   "Carrier_63_G120DControlWord.2" AT %I3510.2 : Bool;   // Bit_02_AUS3_STOP
   "Carrier_63_G120DControlWord.3" AT %I3510.3 : Bool;   // Bit_03_EN
   "Carrier_63_G120DControlWord.4" AT %I3510.4 : Bool;   // Bit_04_EN_RAMP
   "Carrier_63_G120DControlWord.5" AT %I3510.5 : Bool;   // Bit_05_START_RAMP
   "Carrier_63_G120DControlWord.6" AT %I3510.6 : Bool;   // Bit_06_SETPOINT
   "Carrier_63_G120DControlWord.7" AT %I3510.7 : Bool;   // Bit_07_RESET
   "Carrier_63_G120DControlWord.8" AT %I3511.0 : Bool;   // Bit_08_JOG_R
   "Carrier_63_G120DControlWord.9" AT %I3511.1 : Bool;   // Bit_09_JOG_L
   "Carrier_63_G120DControlWord.10" AT %I3511.2 : Bool;   // Bit_10_CONTR_PLC
   "Carrier_63_G120DControlWord.11" AT %I3511.3 : Bool;   // Bit_11_REVERSE
   "Carrier_63_G120DControlWord.12" AT %I3511.4 : Bool;   // Bit_12_BRAKE_RELEASE
   "Carrier_63_G120DControlWord.13" AT %I3511.5 : Bool;   // Bit_13_DDS
   "Carrier_63_G120DControlWord.14" AT %I3511.6 : Bool;   // Bit_14_DO0
   "Carrier_63_G120DControlWord.15" AT %I3511.7 : Bool;   // Bit_15_DO1
   "Carrier_63_G120DStatusWord" AT %IW3512 : Word;   // G120D_ZSW1_STATUS
   "Carrier_63_G120DStatusWord.0" AT %I3512.0 : Bool;   // Bit_00_READY_RUN
   "Carrier_63_G120DStatusWord.1" AT %I3512.1 : Bool;   // Bit_01_READY_ON
   "Carrier_63_G120DStatusWord.2" AT %I3512.2 : Bool;   // Bit_02_ENABLE
   "Carrier_63_G120DStatusWord.3" AT %I3512.3 : Bool;   // Bit_03_FAULT
   "Carrier_63_G120DStatusWord.4" AT %I3512.4 : Bool;   // Bit_04_OFF2
   "Carrier_63_G120DStatusWord.5" AT %I3512.5 : Bool;   // Bit_05_OFF3
   "Carrier_63_G120DStatusWord.6" AT %I3512.6 : Bool;   // Bit_06_LOCK_OUT
   "Carrier_63_G120DStatusWord.7" AT %I3512.7 : Bool;   // Bit_07_WARN
   "Carrier_63_G120DStatusWord.8" AT %I3513.0 : Bool;   // Bit_08_NO_DEVIATION
   "Carrier_63_G120DStatusWord.9" AT %I3513.1 : Bool;   // Bit_09_CONTR_PLC
   "Carrier_63_G120DStatusWord.10" AT %I3513.2 : Bool;   // Bit_10_F_MAX
   "Carrier_63_G120DStatusWord.11" AT %I3513.3 : Bool;   // Bit_11_LIMIT_REACHED
   "Carrier_63_G120DStatusWord.12" AT %I3513.4 : Bool;   // Bit_12_BRAKE_OPEN
   "Carrier_63_G120DStatusWord.13" AT %I3513.5 : Bool;   // Bit_13_NO_OVERTEMP
   "Carrier_63_G120DStatusWord.14" AT %I3513.6 : Bool;   // Bit_14_CW_CCW
   "Carrier_63_G120DStatusWord.15" AT %I3513.7 : Bool;   // Bit_15_OVERL
   "Carrier_63_Slot2_Input" AT %IW3514 : Word;   // SLOT 2 INPUT WORD
   "Carrier_63_CrashDetectSW" AT %I3514.0 : Bool;   // CRASH DETECT SW
   "Carrier_63_SpareSafetyInput(2_1)" AT %I3514.1 : Bool;   // SPARE SAFETY INPUT
   "Carrier_63_SpareSafetyInput(2_2)" AT %I3514.2 : Bool;   // SPARE SAFETY INPUT
   "Carrier_63_SpareSafetyInput(2_3)" AT %I3514.3 : Bool;   // SPARE SAFETY INPUT
   "Carrier_63_SpareSafetyInput(2_4)" AT %I3514.4 : Bool;   // SPARE SAFETY INPUT
   "Carrier_63_SpareSafetyInput(2_5)" AT %I3514.5 : Bool;   // SPARE SAFETY INPUT
   "Carrier_63_SpareSafetyInput(2_6)" AT %I3514.6 : Bool;   // SPARE SAFETY INPUT
   "Carrier_63_SpareSafetyInput(2_7)" AT %I3514.7 : Bool;   // SPARE SAFETY INPUT
   "Carrier_63_Slot3_SafetyOutput" AT %IW3515 : Word;   // SLOT 3 SAFETY OUTPUT WORD
   "Carrier_63_Crash_Detect_OK" AT %I3515.0 : Bool;   // CARRIER CRASH DETECT
   "Carrier_63_SpareSafetyOutput(3_1)" AT %I3515.1 : Bool;   // SPARE SAFETY OUTPUT
   "Carrier_63_SpareSafetyOutput(3_2)" AT %I3515.2 : Bool;   // SPARE SAFETY OUTPUT
   "Carrier_63_SpareSafetyOutput(3_3)" AT %I3515.3 : Bool;   // SPARE SAFETY OUTPUT
   "Carrier_63_SpareSafetyOutput(3_4)" AT %I3515.4 : Bool;   // SPARE SAFETY OUTPUT
   "Carrier_63_SpareSafetyOutput(3_5)" AT %I3515.5 : Bool;   // SPARE SAFETY OUTPUT
   "Carrier_63_SpareSafetyOutput(3_6)" AT %I3515.6 : Bool;   // SPARE SAFETY OUTPUT
   "Carrier_63_SpareSafetyOutput(3_7)" AT %I3515.7 : Bool;   // SPARE SAFETY OUTPUT
   "Carrier_63_Slot4_Input" AT %IW3516 : Word;   // SLOT 4 INPUT WORD
   "Carrier_63_480VPowerOn_MDCB1" AT %I3516.0 : Bool;   // 480 VAC POWER ON MDCB 1
   "Carrier_63_SpareInput(4_1)" AT %I3516.1 : Bool;   // SPARE INPUT
   "Carrier_63_SpareInput(4_2)" AT %I3516.2 : Bool;   // SPARE INPUT
   "Carrier_63_SitopSelectStatus" AT %I3516.3 : Bool;   // SITOP SELECT STATUS
   "Carrier_63_DCsupplyOnPSCB2" AT %I3516.4 : Bool;   // DC SUPPLY ON PSCB 2
   "Carrier_63_SpareInput(4_5)" AT %I3516.5 : Bool;   // SPARE INPUT
   "Carrier_63_SpareInput(4_6)" AT %I3516.6 : Bool;   // SPARE INPUT
   "Carrier_63_SpareInput(4_7)" AT %I3516.7 : Bool;   // SPARE INPUT
   "Carrier_63_PB1_ProdHoldLH" AT %I3517.0 : Bool;   // PB 1 PRODUCTION HOLD LH
   "Carrier_63_PB2_ResetLH" AT %I3517.1 : Bool;   // PB 2 RESET LH
   "Carrier_63_PB3_ProdHoldRH" AT %I3517.2 : Bool;   // PB 3 PRODUCTION HOLD RH
   "Carrier_63_PB4_ResetRH" AT %I3517.3 : Bool;   // PB 4 RESET RH
   "Carrier_63_SpareInput(4_14)" AT %I3517.4 : Bool;   // SPARE INPUT
   "Carrier_63_SpareInput(4_15)" AT %I3517.5 : Bool;   // SPARE INPUT
   "Carrier_63_SpareInput(4_16)" AT %I3517.6 : Bool;   // SPARE INPUT
   "Carrier_63_SpareInput(4_17)" AT %I3517.7 : Bool;   // SPARE INPUT
   "Carrier_63_Slot5_Output" AT %IW3518 : Word;   // SLOT 5 OUTPUT WORD
   "Carrier_63_IRD400_HMI_24VDC_ENABLE" AT %I3518.0 : Bool;   // IRD 400 PANEL HMI 24V DC POWER
   "Carrier_63_FaultLight_LH" AT %I3518.1 : Bool;   // FAULT LIGHT LH
   "Carrier_63_RunLight_LH" AT %I3518.2 : Bool;   // RUN LIGHT LH
   "Carrier_63_FaultLight_RH" AT %I3518.3 : Bool;   // FAULT LIGHT RH
   "Carrier_63_RunLight_RH" AT %I3518.4 : Bool;   // RUN LIGHT RH
   "Carrier_63_SpareOutput(5_5)" AT %I3518.5 : Bool;   // SPARE OUTPUT
   "Carrier_63_SpareOutput(5_6)" AT %I3518.6 : Bool;   // SPARE OUTPUT
   "Carrier_63_SpareOutput(5_7)" AT %I3518.7 : Bool;   // SPARE OUTPUT
   "Carrier_63_ActualSpeed" AT %IW3520 : Word;   // ACTUAL SPEED
   "Carrier_63_CarrierDriveAlarm" AT %IW3522 : Word;   // CARRIER DRIVE ALARM
   "Carrier_63_CarrierDriveWarning" AT %IW3524 : Word;   // CARRIER DRIVE WARNING
   "Carrier_64_Status" AT %IW3550 : Word;   // CARRIER STATUS WORD
   "Carrier_64_Status.0" AT %I3550.0 : Bool;   // HEARTBEAT
   "Carrier_64_Status.1" AT %I3550.1 : Bool;   // MANUAL
   "Carrier_64_Status.2" AT %I3550.2 : Bool;   // IN_AUTO
   "Carrier_64_Status.3" AT %I3550.3 : Bool;   // POSITIONING_COMPLETE
   "Carrier_64_Status.4" AT %I3550.4 : Bool;   // PRODUCTION HOLD
   "Carrier_64_Status.5" AT %I3550.5 : Bool;   // CARRIER MOVING FORWARD
   "Carrier_64_Status.6" AT %I3550.6 : Bool;   // CARRIER MOVING REVERSE
   "Carrier_64_Status.7" AT %I3550.7 : Bool;   // CARRIER FAULT
   "Carrier_64_Status.8" AT %I3551.0 : Bool;   // CRASH DETECT TRIPPED
   "Carrier_64_Status.9" AT %I3551.1 : Bool;
   "Carrier_64_Status.10" AT %I3551.2 : Bool;
   "Carrier_64_Status.11" AT %I3551.3 : Bool;
   "Carrier_64_Status.12" AT %I3551.4 : Bool;
   "Carrier_64_Status.13" AT %I3551.5 : Bool;
   "Carrier_64_Status.14" AT %I3551.6 : Bool;
   "Carrier_64_Status.15" AT %I3551.7 : Bool;
   "Carrier_64_SDCFaultCode" AT %IW3552 : Word;   // SDC FAULT CODE
   "Carrier_64_CarrierPosition" AT %ID3554 : DWord;   // CARRIER POSITION
   "Carrier_64_CarrierNumber" AT %IW3558 : Word;   // CARRIER NUMBER
   "Carrier_64_G120DControlWord" AT %IW3560 : Word;   // G120D_STW1_CONTROL
   "Carrier_64_G120DControlWord.0" AT %I3560.0 : Bool;   // Bit_00_ON
   "Carrier_64_G120DControlWord.1" AT %I3560.1 : Bool;   // Bit_01_AUS2_INH
   "Carrier_64_G120DControlWord.2" AT %I3560.2 : Bool;   // Bit_02_AUS3_STOP
   "Carrier_64_G120DControlWord.3" AT %I3560.3 : Bool;   // Bit_03_EN
   "Carrier_64_G120DControlWord.4" AT %I3560.4 : Bool;   // Bit_04_EN_RAMP
   "Carrier_64_G120DControlWord.5" AT %I3560.5 : Bool;   // Bit_05_START_RAMP
   "Carrier_64_G120DControlWord.6" AT %I3560.6 : Bool;   // Bit_06_SETPOINT
   "Carrier_64_G120DControlWord.7" AT %I3560.7 : Bool;   // Bit_07_RESET
   "Carrier_64_G120DControlWord.8" AT %I3561.0 : Bool;   // Bit_08_JOG_R
   "Carrier_64_G120DControlWord.9" AT %I3561.1 : Bool;   // Bit_09_JOG_L
   "Carrier_64_G120DControlWord.10" AT %I3561.2 : Bool;   // Bit_10_CONTR_PLC
   "Carrier_64_G120DControlWord.11" AT %I3561.3 : Bool;   // Bit_11_REVERSE
   "Carrier_64_G120DControlWord.12" AT %I3561.4 : Bool;   // Bit_12_BRAKE_RELEASE
   "Carrier_64_G120DControlWord.13" AT %I3561.5 : Bool;   // Bit_13_DDS
   "Carrier_64_G120DControlWord.14" AT %I3561.6 : Bool;   // Bit_14_DO0
   "Carrier_64_G120DControlWord.15" AT %I3561.7 : Bool;   // Bit_15_DO1
   "Carrier_64_G120DStatusWord" AT %IW3562 : Word;   // G120D_ZSW1_STATUS
   "Carrier_64_G120DStatusWord.0" AT %I3562.0 : Bool;   // Bit_00_READY_RUN
   "Carrier_64_G120DStatusWord.1" AT %I3562.1 : Bool;   // Bit_01_READY_ON
   "Carrier_64_G120DStatusWord.2" AT %I3562.2 : Bool;   // Bit_02_ENABLE
   "Carrier_64_G120DStatusWord.3" AT %I3562.3 : Bool;   // Bit_03_FAULT
   "Carrier_64_G120DStatusWord.4" AT %I3562.4 : Bool;   // Bit_04_OFF2
   "Carrier_64_G120DStatusWord.5" AT %I3562.5 : Bool;   // Bit_05_OFF3
   "Carrier_64_G120DStatusWord.6" AT %I3562.6 : Bool;   // Bit_06_LOCK_OUT
   "Carrier_64_G120DStatusWord.7" AT %I3562.7 : Bool;   // Bit_07_WARN
   "Carrier_64_G120DStatusWord.8" AT %I3563.0 : Bool;   // Bit_08_NO_DEVIATION
   "Carrier_64_G120DStatusWord.9" AT %I3563.1 : Bool;   // Bit_09_CONTR_PLC
   "Carrier_64_G120DStatusWord.10" AT %I3563.2 : Bool;   // Bit_10_F_MAX
   "Carrier_64_G120DStatusWord.11" AT %I3563.3 : Bool;   // Bit_11_LIMIT_REACHED
   "Carrier_64_G120DStatusWord.12" AT %I3563.4 : Bool;   // Bit_12_BRAKE_OPEN
   "Carrier_64_G120DStatusWord.13" AT %I3563.5 : Bool;   // Bit_13_NO_OVERTEMP
   "Carrier_64_G120DStatusWord.14" AT %I3563.6 : Bool;   // Bit_14_CW_CCW
   "Carrier_64_G120DStatusWord.15" AT %I3563.7 : Bool;   // Bit_15_OVERL
   "Carrier_64_Slot2_Input" AT %IW3564 : Word;   // SLOT 2 INPUT WORD
   "Carrier_64_CrashDetectSW" AT %I3564.0 : Bool;   // CRASH DETECT SW
   "Carrier_64_SpareSafetyInput(2_1)" AT %I3564.1 : Bool;   // SPARE SAFETY INPUT
   "Carrier_64_SpareSafetyInput(2_2)" AT %I3564.2 : Bool;   // SPARE SAFETY INPUT
   "Carrier_64_SpareSafetyInput(2_3)" AT %I3564.3 : Bool;   // SPARE SAFETY INPUT
   "Carrier_64_SpareSafetyInput(2_4)" AT %I3564.4 : Bool;   // SPARE SAFETY INPUT
   "Carrier_64_SpareSafetyInput(2_5)" AT %I3564.5 : Bool;   // SPARE SAFETY INPUT
   "Carrier_64_SpareSafetyInput(2_6)" AT %I3564.6 : Bool;   // SPARE SAFETY INPUT
   "Carrier_64_SpareSafetyInput(2_7)" AT %I3564.7 : Bool;   // SPARE SAFETY INPUT
   "Carrier_64_Slot3_SafetyOutput" AT %IW3565 : Word;   // SLOT 3 SAFETY OUTPUT WORD
   "Carrier_64_Crash_Detect_OK" AT %I3565.0 : Bool;   // CARRIER CRASH DETECT
   "Carrier_64_SpareSafetyOutput(3_1)" AT %I3565.1 : Bool;   // SPARE SAFETY OUTPUT
   "Carrier_64_SpareSafetyOutput(3_2)" AT %I3565.2 : Bool;   // SPARE SAFETY OUTPUT
   "Carrier_64_SpareSafetyOutput(3_3)" AT %I3565.3 : Bool;   // SPARE SAFETY OUTPUT
   "Carrier_64_SpareSafetyOutput(3_4)" AT %I3565.4 : Bool;   // SPARE SAFETY OUTPUT
   "Carrier_64_SpareSafetyOutput(3_5)" AT %I3565.5 : Bool;   // SPARE SAFETY OUTPUT
   "Carrier_64_SpareSafetyOutput(3_6)" AT %I3565.6 : Bool;   // SPARE SAFETY OUTPUT
   "Carrier_64_SpareSafetyOutput(3_7)" AT %I3565.7 : Bool;   // SPARE SAFETY OUTPUT
   "Carrier_64_Slot4_Input" AT %IW3566 : Word;   // SLOT 4 INPUT WORD
   "Carrier_64_480VPowerOn_MDCB1" AT %I3566.0 : Bool;   // 480 VAC POWER ON MDCB 1
   "Carrier_64_SpareInput(4_1)" AT %I3566.1 : Bool;   // SPARE INPUT
   "Carrier_64_SpareInput(4_2)" AT %I3566.2 : Bool;   // SPARE INPUT
   "Carrier_64_SitopSelectStatus" AT %I3566.3 : Bool;   // SITOP SELECT STATUS
   "Carrier_64_DCsupplyOnPSCB2" AT %I3566.4 : Bool;   // DC SUPPLY ON PSCB 2
   "Carrier_64_SpareInput(4_5)" AT %I3566.5 : Bool;   // SPARE INPUT
   "Carrier_64_SpareInput(4_6)" AT %I3566.6 : Bool;   // SPARE INPUT
   "Carrier_64_SpareInput(4_7)" AT %I3566.7 : Bool;   // SPARE INPUT
   "Carrier_64_PB1_ProdHoldLH" AT %I3567.0 : Bool;   // PB 1 PRODUCTION HOLD LH
   "Carrier_64_PB2_ResetLH" AT %I3567.1 : Bool;   // PB 2 RESET LH
   "Carrier_64_PB3_ProdHoldRH" AT %I3567.2 : Bool;   // PB 3 PRODUCTION HOLD RH
   "Carrier_64_PB4_ResetRH" AT %I3567.3 : Bool;   // PB 4 RESET RH
   "Carrier_64_SpareInput(4_14)" AT %I3567.4 : Bool;   // SPARE INPUT
   "Carrier_64_SpareInput(4_15)" AT %I3567.5 : Bool;   // SPARE INPUT
   "Carrier_64_SpareInput(4_16)" AT %I3567.6 : Bool;   // SPARE INPUT
   "Carrier_64_SpareInput(4_17)" AT %I3567.7 : Bool;   // SPARE INPUT
   "Carrier_64_Slot5_Output" AT %IW3568 : Word;   // SLOT 5 OUTPUT WORD
   "Carrier_64_IRD400_HMI_24VDC_ENABLE" AT %I3568.0 : Bool;   // IRD 400 PANEL HMI 24V DC POWER
   "Carrier_64_FaultLight_LH" AT %I3568.1 : Bool;   // FAULT LIGHT LH
   "Carrier_64_RunLight_LH" AT %I3568.2 : Bool;   // RUN LIGHT LH
   "Carrier_64_FaultLight_RH" AT %I3568.3 : Bool;   // FAULT LIGHT RH
   "Carrier_64_RunLight_RH" AT %I3568.4 : Bool;   // RUN LIGHT RH
   "Carrier_64_SpareOutput(5_5)" AT %I3568.5 : Bool;   // SPARE OUTPUT
   "Carrier_64_SpareOutput(5_6)" AT %I3568.6 : Bool;   // SPARE OUTPUT
   "Carrier_64_SpareOutput(5_7)" AT %I3568.7 : Bool;   // SPARE OUTPUT
   "Carrier_64_ActualSpeed" AT %IW3570 : Word;   // ACTUAL SPEED
   "Carrier_64_CarrierDriveAlarm" AT %IW3572 : Word;   // CARRIER DRIVE ALARM
   "Carrier_64_CarrierDriveWarning" AT %IW3574 : Word;   // CARRIER DRIVE WARNING
   "Carrier_65_Status" AT %IW3600 : Word;   // CARRIER STATUS WORD
   "Carrier_65_Status.0" AT %I3600.0 : Bool;   // HEARTBEAT
   "Carrier_65_Status.1" AT %I3600.1 : Bool;   // MANUAL
   "Carrier_65_Status.2" AT %I3600.2 : Bool;   // IN_AUTO
   "Carrier_65_Status.3" AT %I3600.3 : Bool;   // POSITIONING_COMPLETE
   "Carrier_65_Status.4" AT %I3600.4 : Bool;   // PRODUCTION HOLD
   "Carrier_65_Status.5" AT %I3600.5 : Bool;   // CARRIER MOVING FORWARD
   "Carrier_65_Status.6" AT %I3600.6 : Bool;   // CARRIER MOVING REVERSE
   "Carrier_65_Status.7" AT %I3600.7 : Bool;   // CARRIER FAULT
   "Carrier_65_Status.8" AT %I3601.0 : Bool;   // CRASH DETECT TRIPPED
   "Carrier_65_Status.9" AT %I3601.1 : Bool;
   "Carrier_65_Status.10" AT %I3601.2 : Bool;
   "Carrier_65_Status.11" AT %I3601.3 : Bool;
   "Carrier_65_Status.12" AT %I3601.4 : Bool;
   "Carrier_65_Status.13" AT %I3601.5 : Bool;
   "Carrier_65_Status.14" AT %I3601.6 : Bool;
   "Carrier_65_Status.15" AT %I3601.7 : Bool;
   "Carrier_65_SDCFaultCode" AT %IW3602 : Word;   // SDC FAULT CODE
   "Carrier_65_CarrierPosition" AT %ID3604 : DWord;   // CARRIER POSITION
   "Carrier_65_CarrierNumber" AT %IW3608 : Word;   // CARRIER NUMBER
   "Carrier_65_G120DControlWord" AT %IW3600 : Word;   // G120D_STW1_CONTROL
   "Carrier_65_G120DControlWord.0" AT %I3600.0 : Bool;   // Bit_00_ON
   "Carrier_65_G120DControlWord.1" AT %I3600.1 : Bool;   // Bit_01_AUS2_INH
   "Carrier_65_G120DControlWord.2" AT %I3600.2 : Bool;   // Bit_02_AUS3_STOP
   "Carrier_65_G120DControlWord.3" AT %I3600.3 : Bool;   // Bit_03_EN
   "Carrier_65_G120DControlWord.4" AT %I3600.4 : Bool;   // Bit_04_EN_RAMP
   "Carrier_65_G120DControlWord.5" AT %I3600.5 : Bool;   // Bit_05_START_RAMP
   "Carrier_65_G120DControlWord.6" AT %I3600.6 : Bool;   // Bit_06_SETPOINT
   "Carrier_65_G120DControlWord.7" AT %I3600.7 : Bool;   // Bit_07_RESET
   "Carrier_65_G120DControlWord.8" AT %I3601.0 : Bool;   // Bit_08_JOG_R
   "Carrier_65_G120DControlWord.9" AT %I3601.1 : Bool;   // Bit_09_JOG_L
   "Carrier_65_G120DControlWord.10" AT %I3601.2 : Bool;   // Bit_10_CONTR_PLC
   "Carrier_65_G120DControlWord.11" AT %I3601.3 : Bool;   // Bit_11_REVERSE
   "Carrier_65_G120DControlWord.12" AT %I3601.4 : Bool;   // Bit_12_BRAKE_RELEASE
   "Carrier_65_G120DControlWord.13" AT %I3601.5 : Bool;   // Bit_13_DDS
   "Carrier_65_G120DControlWord.14" AT %I3601.6 : Bool;   // Bit_14_DO0
   "Carrier_65_G120DControlWord.15" AT %I3601.7 : Bool;   // Bit_15_DO1
   "Carrier_65_G120DStatusWord" AT %IW3602 : Word;   // G120D_ZSW1_STATUS
   "Carrier_65_G120DStatusWord.0" AT %I3602.0 : Bool;   // Bit_00_READY_RUN
   "Carrier_65_G120DStatusWord.1" AT %I3602.1 : Bool;   // Bit_01_READY_ON
   "Carrier_65_G120DStatusWord.2" AT %I3602.2 : Bool;   // Bit_02_ENABLE
   "Carrier_65_G120DStatusWord.3" AT %I3602.3 : Bool;   // Bit_03_FAULT
   "Carrier_65_G120DStatusWord.4" AT %I3602.4 : Bool;   // Bit_04_OFF2
   "Carrier_65_G120DStatusWord.5" AT %I3602.5 : Bool;   // Bit_05_OFF3
   "Carrier_65_G120DStatusWord.6" AT %I3602.6 : Bool;   // Bit_06_LOCK_OUT
   "Carrier_65_G120DStatusWord.7" AT %I3602.7 : Bool;   // Bit_07_WARN
   "Carrier_65_G120DStatusWord.8" AT %I3603.0 : Bool;   // Bit_08_NO_DEVIATION
   "Carrier_65_G120DStatusWord.9" AT %I3603.1 : Bool;   // Bit_09_CONTR_PLC
   "Carrier_65_G120DStatusWord.10" AT %I3603.2 : Bool;   // Bit_10_F_MAX
   "Carrier_65_G120DStatusWord.11" AT %I3603.3 : Bool;   // Bit_11_LIMIT_REACHED
   "Carrier_65_G120DStatusWord.12" AT %I3603.4 : Bool;   // Bit_12_BRAKE_OPEN
   "Carrier_65_G120DStatusWord.13" AT %I3603.5 : Bool;   // Bit_13_NO_OVERTEMP
   "Carrier_65_G120DStatusWord.14" AT %I3603.6 : Bool;   // Bit_14_CW_CCW
   "Carrier_65_G120DStatusWord.15" AT %I3603.7 : Bool;   // Bit_15_OVERL
   "Carrier_65_Slot2_Input" AT %IW3604 : Word;   // SLOT 2 INPUT WORD
   "Carrier_65_CrashDetectSW" AT %I3604.0 : Bool;   // CRASH DETECT SW
   "Carrier_65_SpareSafetyInput(2_1)" AT %I3604.1 : Bool;   // SPARE SAFETY INPUT
   "Carrier_65_SpareSafetyInput(2_2)" AT %I3604.2 : Bool;   // SPARE SAFETY INPUT
   "Carrier_65_SpareSafetyInput(2_3)" AT %I3604.3 : Bool;   // SPARE SAFETY INPUT
   "Carrier_65_SpareSafetyInput(2_4)" AT %I3604.4 : Bool;   // SPARE SAFETY INPUT
   "Carrier_65_SpareSafetyInput(2_5)" AT %I3604.5 : Bool;   // SPARE SAFETY INPUT
   "Carrier_65_SpareSafetyInput(2_6)" AT %I3604.6 : Bool;   // SPARE SAFETY INPUT
   "Carrier_65_SpareSafetyInput(2_7)" AT %I3604.7 : Bool;   // SPARE SAFETY INPUT
   "Carrier_65_Slot3_SafetyOutput" AT %IW3605 : Word;   // SLOT 3 SAFETY OUTPUT WORD
   "Carrier_65_Crash_Detect_OK" AT %I3605.0 : Bool;   // CARRIER CRASH DETECT
   "Carrier_65_SpareSafetyOutput(3_1)" AT %I3605.1 : Bool;   // SPARE SAFETY OUTPUT
   "Carrier_65_SpareSafetyOutput(3_2)" AT %I3605.2 : Bool;   // SPARE SAFETY OUTPUT
   "Carrier_65_SpareSafetyOutput(3_3)" AT %I3605.3 : Bool;   // SPARE SAFETY OUTPUT
   "Carrier_65_SpareSafetyOutput(3_4)" AT %I3605.4 : Bool;   // SPARE SAFETY OUTPUT
   "Carrier_65_SpareSafetyOutput(3_5)" AT %I3605.5 : Bool;   // SPARE SAFETY OUTPUT
   "Carrier_65_SpareSafetyOutput(3_6)" AT %I3605.6 : Bool;   // SPARE SAFETY OUTPUT
   "Carrier_65_SpareSafetyOutput(3_7)" AT %I3605.7 : Bool;   // SPARE SAFETY OUTPUT
   "Carrier_65_Slot4_Input" AT %IW3606 : Word;   // SLOT 4 INPUT WORD
   "Carrier_65_480VPowerOn_MDCB1" AT %I3606.0 : Bool;   // 480 VAC POWER ON MDCB 1
   "Carrier_65_SpareInput(4_1)" AT %I3606.1 : Bool;   // SPARE INPUT
   "Carrier_65_SpareInput(4_2)" AT %I3606.2 : Bool;   // SPARE INPUT
   "Carrier_65_SitopSelectStatus" AT %I3606.3 : Bool;   // SITOP SELECT STATUS
   "Carrier_65_DCsupplyOnPSCB2" AT %I3606.4 : Bool;   // DC SUPPLY ON PSCB 2
   "Carrier_65_SpareInput(4_5)" AT %I3606.5 : Bool;   // SPARE INPUT
   "Carrier_65_SpareInput(4_6)" AT %I3606.6 : Bool;   // SPARE INPUT
   "Carrier_65_SpareInput(4_7)" AT %I3606.7 : Bool;   // SPARE INPUT
   "Carrier_65_PB1_ProdHoldLH" AT %I3607.0 : Bool;   // PB 1 PRODUCTION HOLD LH
   "Carrier_65_PB2_ResetLH" AT %I3607.1 : Bool;   // PB 2 RESET LH
   "Carrier_65_PB3_ProdHoldRH" AT %I3607.2 : Bool;   // PB 3 PRODUCTION HOLD RH
   "Carrier_65_PB4_ResetRH" AT %I3607.3 : Bool;   // PB 4 RESET RH
   "Carrier_65_SpareInput(4_14)" AT %I3607.4 : Bool;   // SPARE INPUT
   "Carrier_65_SpareInput(4_15)" AT %I3607.5 : Bool;   // SPARE INPUT
   "Carrier_65_SpareInput(4_16)" AT %I3607.6 : Bool;   // SPARE INPUT
   "Carrier_65_SpareInput(4_17)" AT %I3607.7 : Bool;   // SPARE INPUT
   "Carrier_65_Slot5_Output" AT %IW3608 : Word;   // SLOT 5 OUTPUT WORD
   "Carrier_65_IRD400_HMI_24VDC_ENABLE" AT %I3608.0 : Bool;   // IRD 400 PANEL HMI 24V DC POWER
   "Carrier_65_FaultLight_LH" AT %I3608.1 : Bool;   // FAULT LIGHT LH
   "Carrier_65_RunLight_LH" AT %I3608.2 : Bool;   // RUN LIGHT LH
   "Carrier_65_FaultLight_RH" AT %I3608.3 : Bool;   // FAULT LIGHT RH
   "Carrier_65_RunLight_RH" AT %I3608.4 : Bool;   // RUN LIGHT RH
   "Carrier_65_SpareOutput(5_5)" AT %I3608.5 : Bool;   // SPARE OUTPUT
   "Carrier_65_SpareOutput(5_6)" AT %I3608.6 : Bool;   // SPARE OUTPUT
   "Carrier_65_SpareOutput(5_7)" AT %I3608.7 : Bool;   // SPARE OUTPUT
   "Carrier_65_ActualSpeed" AT %IW3620 : Word;   // ACTUAL SPEED
   "Carrier_65_CarrierDriveAlarm" AT %IW3622 : Word;   // CARRIER DRIVE ALARM
   "Carrier_65_CarrierDriveWarning" AT %IW3624 : Word;   // CARRIER DRIVE WARNING
   "Carrier_66_Status" AT %IW3650 : Word;   // CARRIER STATUS WORD
   "Carrier_66_Status.0" AT %I3650.0 : Bool;   // HEARTBEAT
   "Carrier_66_Status.1" AT %I3650.1 : Bool;   // MANUAL
   "Carrier_66_Status.2" AT %I3650.2 : Bool;   // IN_AUTO
   "Carrier_66_Status.3" AT %I3650.3 : Bool;   // POSITIONING_COMPLETE
   "Carrier_66_Status.4" AT %I3650.4 : Bool;   // PRODUCTION HOLD
   "Carrier_66_Status.5" AT %I3650.5 : Bool;   // CARRIER MOVING FORWARD
   "Carrier_66_Status.6" AT %I3650.6 : Bool;   // CARRIER MOVING REVERSE
   "Carrier_66_Status.7" AT %I3650.7 : Bool;   // CARRIER FAULT
   "Carrier_66_Status.8" AT %I3651.0 : Bool;   // CRASH DETECT TRIPPED
   "Carrier_66_Status.9" AT %I3651.1 : Bool;
   "Carrier_66_Status.10" AT %I3651.2 : Bool;
   "Carrier_66_Status.11" AT %I3651.3 : Bool;
   "Carrier_66_Status.12" AT %I3651.4 : Bool;
   "Carrier_66_Status.13" AT %I3651.5 : Bool;
   "Carrier_66_Status.14" AT %I3651.6 : Bool;
   "Carrier_66_Status.15" AT %I3651.7 : Bool;
   "Carrier_66_SDCFaultCode" AT %IW3652 : Word;   // SDC FAULT CODE
   "Carrier_66_CarrierPosition" AT %ID3654 : DWord;   // CARRIER POSITION
   "Carrier_66_CarrierNumber" AT %IW3658 : Word;   // CARRIER NUMBER
   "Carrier_66_G120DControlWord" AT %IW3660 : Word;   // G120D_STW1_CONTROL
   "Carrier_66_G120DControlWord.0" AT %I3660.0 : Bool;   // Bit_00_ON
   "Carrier_66_G120DControlWord.1" AT %I3660.1 : Bool;   // Bit_01_AUS2_INH
   "Carrier_66_G120DControlWord.2" AT %I3660.2 : Bool;   // Bit_02_AUS3_STOP
   "Carrier_66_G120DControlWord.3" AT %I3660.3 : Bool;   // Bit_03_EN
   "Carrier_66_G120DControlWord.4" AT %I3660.4 : Bool;   // Bit_04_EN_RAMP
   "Carrier_66_G120DControlWord.5" AT %I3660.5 : Bool;   // Bit_05_START_RAMP
   "Carrier_66_G120DControlWord.6" AT %I3660.6 : Bool;   // Bit_06_SETPOINT
   "Carrier_66_G120DControlWord.7" AT %I3660.7 : Bool;   // Bit_07_RESET
   "Carrier_66_G120DControlWord.8" AT %I3661.0 : Bool;   // Bit_08_JOG_R
   "Carrier_66_G120DControlWord.9" AT %I3661.1 : Bool;   // Bit_09_JOG_L
   "Carrier_66_G120DControlWord.10" AT %I3661.2 : Bool;   // Bit_10_CONTR_PLC
   "Carrier_66_G120DControlWord.11" AT %I3661.3 : Bool;   // Bit_11_REVERSE
   "Carrier_66_G120DControlWord.12" AT %I3661.4 : Bool;   // Bit_12_BRAKE_RELEASE
   "Carrier_66_G120DControlWord.13" AT %I3661.5 : Bool;   // Bit_13_DDS
   "Carrier_66_G120DControlWord.14" AT %I3661.6 : Bool;   // Bit_14_DO0
   "Carrier_66_G120DControlWord.15" AT %I3661.7 : Bool;   // Bit_15_DO1
   "Carrier_66_G120DStatusWord" AT %IW3662 : Word;   // G120D_ZSW1_STATUS
   "Carrier_66_G120DStatusWord.0" AT %I3662.0 : Bool;   // Bit_00_READY_RUN
   "Carrier_66_G120DStatusWord.1" AT %I3662.1 : Bool;   // Bit_01_READY_ON
   "Carrier_66_G120DStatusWord.2" AT %I3662.2 : Bool;   // Bit_02_ENABLE
   "Carrier_66_G120DStatusWord.3" AT %I3662.3 : Bool;   // Bit_03_FAULT
   "Carrier_66_G120DStatusWord.4" AT %I3662.4 : Bool;   // Bit_04_OFF2
   "Carrier_66_G120DStatusWord.5" AT %I3662.5 : Bool;   // Bit_05_OFF3
   "Carrier_66_G120DStatusWord.6" AT %I3662.6 : Bool;   // Bit_06_LOCK_OUT
   "Carrier_66_G120DStatusWord.7" AT %I3662.7 : Bool;   // Bit_07_WARN
   "Carrier_66_G120DStatusWord.8" AT %I3663.0 : Bool;   // Bit_08_NO_DEVIATION
   "Carrier_66_G120DStatusWord.9" AT %I3663.1 : Bool;   // Bit_09_CONTR_PLC
   "Carrier_66_G120DStatusWord.10" AT %I3663.2 : Bool;   // Bit_10_F_MAX
   "Carrier_66_G120DStatusWord.11" AT %I3663.3 : Bool;   // Bit_11_LIMIT_REACHED
   "Carrier_66_G120DStatusWord.12" AT %I3663.4 : Bool;   // Bit_12_BRAKE_OPEN
   "Carrier_66_G120DStatusWord.13" AT %I3663.5 : Bool;   // Bit_13_NO_OVERTEMP
   "Carrier_66_G120DStatusWord.14" AT %I3663.6 : Bool;   // Bit_14_CW_CCW
   "Carrier_66_G120DStatusWord.15" AT %I3663.7 : Bool;   // Bit_15_OVERL
   "Carrier_66_Slot2_Input" AT %IW3664 : Word;   // SLOT 2 INPUT WORD
   "Carrier_66_CrashDetectSW" AT %I3664.0 : Bool;   // CRASH DETECT SW
   "Carrier_66_SpareSafetyInput(2_1)" AT %I3664.1 : Bool;   // SPARE SAFETY INPUT
   "Carrier_66_SpareSafetyInput(2_2)" AT %I3664.2 : Bool;   // SPARE SAFETY INPUT
   "Carrier_66_SpareSafetyInput(2_3)" AT %I3664.3 : Bool;   // SPARE SAFETY INPUT
   "Carrier_66_SpareSafetyInput(2_4)" AT %I3664.4 : Bool;   // SPARE SAFETY INPUT
   "Carrier_66_SpareSafetyInput(2_5)" AT %I3664.5 : Bool;   // SPARE SAFETY INPUT
   "Carrier_66_SpareSafetyInput(2_6)" AT %I3664.6 : Bool;   // SPARE SAFETY INPUT
   "Carrier_66_SpareSafetyInput(2_7)" AT %I3664.7 : Bool;   // SPARE SAFETY INPUT
   "Carrier_66_Slot3_SafetyOutput" AT %IW3665 : Word;   // SLOT 3 SAFETY OUTPUT WORD
   "Carrier_66_Crash_Detect_OK" AT %I3665.0 : Bool;   // CARRIER CRASH DETECT
   "Carrier_66_SpareSafetyOutput(3_1)" AT %I3665.1 : Bool;   // SPARE SAFETY OUTPUT
   "Carrier_66_SpareSafetyOutput(3_2)" AT %I3665.2 : Bool;   // SPARE SAFETY OUTPUT
   "Carrier_66_SpareSafetyOutput(3_3)" AT %I3665.3 : Bool;   // SPARE SAFETY OUTPUT
   "Carrier_66_SpareSafetyOutput(3_4)" AT %I3665.4 : Bool;   // SPARE SAFETY OUTPUT
   "Carrier_66_SpareSafetyOutput(3_5)" AT %I3665.5 : Bool;   // SPARE SAFETY OUTPUT
   "Carrier_66_SpareSafetyOutput(3_6)" AT %I3665.6 : Bool;   // SPARE SAFETY OUTPUT
   "Carrier_66_SpareSafetyOutput(3_7)" AT %I3665.7 : Bool;   // SPARE SAFETY OUTPUT
   "Carrier_66_Slot4_Input" AT %IW3666 : Word;   // SLOT 4 INPUT WORD
   "Carrier_66_480VPowerOn_MDCB1" AT %I3666.0 : Bool;   // 480 VAC POWER ON MDCB 1
   "Carrier_66_SpareInput(4_1)" AT %I3666.1 : Bool;   // SPARE INPUT
   "Carrier_66_SpareInput(4_2)" AT %I3666.2 : Bool;   // SPARE INPUT
   "Carrier_66_SitopSelectStatus" AT %I3666.3 : Bool;   // SITOP SELECT STATUS
   "Carrier_66_DCsupplyOnPSCB2" AT %I3666.4 : Bool;   // DC SUPPLY ON PSCB 2
   "Carrier_66_SpareInput(4_5)" AT %I3666.5 : Bool;   // SPARE INPUT
   "Carrier_66_SpareInput(4_6)" AT %I3666.6 : Bool;   // SPARE INPUT
   "Carrier_66_SpareInput(4_7)" AT %I3666.7 : Bool;   // SPARE INPUT
   "Carrier_66_PB1_ProdHoldLH" AT %I3667.0 : Bool;   // PB 1 PRODUCTION HOLD LH
   "Carrier_66_PB2_ResetLH" AT %I3667.1 : Bool;   // PB 2 RESET LH
   "Carrier_66_PB3_ProdHoldRH" AT %I3667.2 : Bool;   // PB 3 PRODUCTION HOLD RH
   "Carrier_66_PB4_ResetRH" AT %I3667.3 : Bool;   // PB 4 RESET RH
   "Carrier_66_SpareInput(4_14)" AT %I3667.4 : Bool;   // SPARE INPUT
   "Carrier_66_SpareInput(4_15)" AT %I3667.5 : Bool;   // SPARE INPUT
   "Carrier_66_SpareInput(4_16)" AT %I3667.6 : Bool;   // SPARE INPUT
   "Carrier_66_SpareInput(4_17)" AT %I3667.7 : Bool;   // SPARE INPUT
   "Carrier_66_Slot5_Output" AT %IW3668 : Word;   // SLOT 5 OUTPUT WORD
   "Carrier_66_IRD400_HMI_24VDC_ENABLE" AT %I3668.0 : Bool;   // IRD 400 PANEL HMI 24V DC POWER
   "Carrier_66_FaultLight_LH" AT %I3668.1 : Bool;   // FAULT LIGHT LH
   "Carrier_66_RunLight_LH" AT %I3668.2 : Bool;   // RUN LIGHT LH
   "Carrier_66_FaultLight_RH" AT %I3668.3 : Bool;   // FAULT LIGHT RH
   "Carrier_66_RunLight_RH" AT %I3668.4 : Bool;   // RUN LIGHT RH
   "Carrier_66_SpareOutput(5_5)" AT %I3668.5 : Bool;   // SPARE OUTPUT
   "Carrier_66_SpareOutput(5_6)" AT %I3668.6 : Bool;   // SPARE OUTPUT
   "Carrier_66_SpareOutput(5_7)" AT %I3668.7 : Bool;   // SPARE OUTPUT
   "Carrier_66_ActualSpeed" AT %IW3670 : Word;   // ACTUAL SPEED
   "Carrier_66_CarrierDriveAlarm" AT %IW3672 : Word;   // CARRIER DRIVE ALARM
   "Carrier_66_CarrierDriveWarning" AT %IW3674 : Word;   // CARRIER DRIVE WARNING
   "Carrier_67_Status" AT %IW3700 : Word;   // CARRIER STATUS WORD
   "Carrier_67_Status.0" AT %I3700.0 : Bool;   // HEARTBEAT
   "Carrier_67_Status.1" AT %I3700.1 : Bool;   // MANUAL
   "Carrier_67_Status.2" AT %I3700.2 : Bool;   // IN_AUTO
   "Carrier_67_Status.3" AT %I3700.3 : Bool;   // POSITIONING_COMPLETE
   "Carrier_67_Status.4" AT %I3700.4 : Bool;   // PRODUCTION HOLD
   "Carrier_67_Status.5" AT %I3700.5 : Bool;   // CARRIER MOVING FORWARD
   "Carrier_67_Status.6" AT %I3700.6 : Bool;   // CARRIER MOVING REVERSE
   "Carrier_67_Status.7" AT %I3700.7 : Bool;   // CARRIER FAULT
   "Carrier_67_Status.8" AT %I3701.0 : Bool;   // CRASH DETECT TRIPPED
   "Carrier_67_Status.9" AT %I3701.1 : Bool;
   "Carrier_67_Status.10" AT %I3701.2 : Bool;
   "Carrier_67_Status.11" AT %I3701.3 : Bool;
   "Carrier_67_Status.12" AT %I3701.4 : Bool;
   "Carrier_67_Status.13" AT %I3701.5 : Bool;
   "Carrier_67_Status.14" AT %I3701.6 : Bool;
   "Carrier_67_Status.15" AT %I3701.7 : Bool;
   "Carrier_67_SDCFaultCode" AT %IW3702 : Word;   // SDC FAULT CODE
   "Carrier_67_CarrierPosition" AT %ID3704 : DWord;   // CARRIER POSITION
   "Carrier_67_CarrierNumber" AT %IW3708 : Word;   // CARRIER NUMBER
   "Carrier_67_G120DControlWord" AT %IW3710 : Word;   // G120D_STW1_CONTROL
   "Carrier_67_G120DControlWord.0" AT %I3710.0 : Bool;   // Bit_00_ON
   "Carrier_67_G120DControlWord.1" AT %I3710.1 : Bool;   // Bit_01_AUS2_INH
   "Carrier_67_G120DControlWord.2" AT %I3710.2 : Bool;   // Bit_02_AUS3_STOP
   "Carrier_67_G120DControlWord.3" AT %I3710.3 : Bool;   // Bit_03_EN
   "Carrier_67_G120DControlWord.4" AT %I3710.4 : Bool;   // Bit_04_EN_RAMP
   "Carrier_67_G120DControlWord.5" AT %I3710.5 : Bool;   // Bit_05_START_RAMP
   "Carrier_67_G120DControlWord.6" AT %I3710.6 : Bool;   // Bit_06_SETPOINT
   "Carrier_67_G120DControlWord.7" AT %I3710.7 : Bool;   // Bit_07_RESET
   "Carrier_67_G120DControlWord.8" AT %I3711.0 : Bool;   // Bit_08_JOG_R
   "Carrier_67_G120DControlWord.9" AT %I3711.1 : Bool;   // Bit_09_JOG_L
   "Carrier_67_G120DControlWord.10" AT %I3711.2 : Bool;   // Bit_10_CONTR_PLC
   "Carrier_67_G120DControlWord.11" AT %I3711.3 : Bool;   // Bit_11_REVERSE
   "Carrier_67_G120DControlWord.12" AT %I3711.4 : Bool;   // Bit_12_BRAKE_RELEASE
   "Carrier_67_G120DControlWord.13" AT %I3711.5 : Bool;   // Bit_13_DDS
   "Carrier_67_G120DControlWord.14" AT %I3711.6 : Bool;   // Bit_14_DO0
   "Carrier_67_G120DControlWord.15" AT %I3711.7 : Bool;   // Bit_15_DO1
   "Carrier_67_G120DStatusWord" AT %IW3712 : Word;   // G120D_ZSW1_STATUS
   "Carrier_67_G120DStatusWord.0" AT %I3712.0 : Bool;   // Bit_00_READY_RUN
   "Carrier_67_G120DStatusWord.1" AT %I3712.1 : Bool;   // Bit_01_READY_ON
   "Carrier_67_G120DStatusWord.2" AT %I3712.2 : Bool;   // Bit_02_ENABLE
   "Carrier_67_G120DStatusWord.3" AT %I3712.3 : Bool;   // Bit_03_FAULT
   "Carrier_67_G120DStatusWord.4" AT %I3712.4 : Bool;   // Bit_04_OFF2
   "Carrier_67_G120DStatusWord.5" AT %I3712.5 : Bool;   // Bit_05_OFF3
   "Carrier_67_G120DStatusWord.6" AT %I3712.6 : Bool;   // Bit_06_LOCK_OUT
   "Carrier_67_G120DStatusWord.7" AT %I3712.7 : Bool;   // Bit_07_WARN
   "Carrier_67_G120DStatusWord.8" AT %I3713.0 : Bool;   // Bit_08_NO_DEVIATION
   "Carrier_67_G120DStatusWord.9" AT %I3713.1 : Bool;   // Bit_09_CONTR_PLC
   "Carrier_67_G120DStatusWord.10" AT %I3713.2 : Bool;   // Bit_10_F_MAX
   "Carrier_67_G120DStatusWord.11" AT %I3713.3 : Bool;   // Bit_11_LIMIT_REACHED
   "Carrier_67_G120DStatusWord.12" AT %I3713.4 : Bool;   // Bit_12_BRAKE_OPEN
   "Carrier_67_G120DStatusWord.13" AT %I3713.5 : Bool;   // Bit_13_NO_OVERTEMP
   "Carrier_67_G120DStatusWord.14" AT %I3713.6 : Bool;   // Bit_14_CW_CCW
   "Carrier_67_G120DStatusWord.15" AT %I3713.7 : Bool;   // Bit_15_OVERL
   "Carrier_67_Slot2_Input" AT %IW3714 : Word;   // SLOT 2 INPUT WORD
   "Carrier_67_CrashDetectSW" AT %I3714.0 : Bool;   // CRASH DETECT SW
   "Carrier_67_SpareSafetyInput(2_1)" AT %I3714.1 : Bool;   // SPARE SAFETY INPUT
   "Carrier_67_SpareSafetyInput(2_2)" AT %I3714.2 : Bool;   // SPARE SAFETY INPUT
   "Carrier_67_SpareSafetyInput(2_3)" AT %I3714.3 : Bool;   // SPARE SAFETY INPUT
   "Carrier_67_SpareSafetyInput(2_4)" AT %I3714.4 : Bool;   // SPARE SAFETY INPUT
   "Carrier_67_SpareSafetyInput(2_5)" AT %I3714.5 : Bool;   // SPARE SAFETY INPUT
   "Carrier_67_SpareSafetyInput(2_6)" AT %I3714.6 : Bool;   // SPARE SAFETY INPUT
   "Carrier_67_SpareSafetyInput(2_7)" AT %I3714.7 : Bool;   // SPARE SAFETY INPUT
   "Carrier_67_Slot3_SafetyOutput" AT %IW3715 : Word;   // SLOT 3 SAFETY OUTPUT WORD
   "Carrier_67_Crash_Detect_OK" AT %I3715.0 : Bool;   // CARRIER CRASH DETECT
   "Carrier_67_SpareSafetyOutput(3_1)" AT %I3715.1 : Bool;   // SPARE SAFETY OUTPUT
   "Carrier_67_SpareSafetyOutput(3_2)" AT %I3715.2 : Bool;   // SPARE SAFETY OUTPUT
   "Carrier_67_SpareSafetyOutput(3_3)" AT %I3715.3 : Bool;   // SPARE SAFETY OUTPUT
   "Carrier_67_SpareSafetyOutput(3_4)" AT %I3715.4 : Bool;   // SPARE SAFETY OUTPUT
   "Carrier_67_SpareSafetyOutput(3_5)" AT %I3715.5 : Bool;   // SPARE SAFETY OUTPUT
   "Carrier_67_SpareSafetyOutput(3_6)" AT %I3715.6 : Bool;   // SPARE SAFETY OUTPUT
   "Carrier_67_SpareSafetyOutput(3_7)" AT %I3715.7 : Bool;   // SPARE SAFETY OUTPUT
   "Carrier_67_Slot4_Input" AT %IW3716 : Word;   // SLOT 4 INPUT WORD
   "Carrier_67_480VPowerOn_MDCB1" AT %I3716.0 : Bool;   // 480 VAC POWER ON MDCB 1
   "Carrier_67_SpareInput(4_1)" AT %I3716.1 : Bool;   // SPARE INPUT
   "Carrier_67_SpareInput(4_2)" AT %I3716.2 : Bool;   // SPARE INPUT
